VERSION : 1.8
// Fehlerliste:
// Nr.(HEX)     Bedeutung:          
// -------------------------------------------------------------------------------
//  00          Kein Fehler
//  01          Lesen/ Schreiben nicht möglich, kein Codeträger im Bereich des 
//              Schreib-/ Lesekopfes
//  02          Fehler beim Lesen
//  03          Codeträger wurde während des Lesens aus dem Bereich des Schreib-/
//              Lesekopfes entfernt
//  04          Fehler beim Schreiben
//  05          Codeträger wurde während des Schreibens aus dem Bereich des
//              Schreib-/ Lesekopfes entfernt
//  06          Zugriffsfehler auf den Speicher
//  07          AV-Bit gesetzt, aber Befehlskennung fehlt oder ist ungültig.
//              oder: Anzahl Byte ist 00
//  09          Kabelbruch Schreib-/ Lesekopf oder Kopf nicht angeschlossen
//  0F          Inhalt der 1. und 2. Bitleiste sind ungleich
//  10          Startadresse + Anzahl byte > Speicherbereich in Initialisierung
//              angegeben
//  11          Ungültige max. Anzahl Schreibzyklen in Initialisierung angegeben
//  12          Ungültige Speichergröße in Initialisierung angegeben
//  13          Ungültige Größe des Speicherbereichs in Initialisierung angegeben
//  14          Ungültige max. Anzahl Schreibzyklen
//  15          Falscher Codeträger-Typ in Initialisierung angegeben
//  16          Max. Anzahl von 2 kByte überschritten
//  17          Codeträger falsch initialisiert (Vergleich mit Vorgabedaten über
//              Befehlskennung 09 Hex bringt keine Übereinstimmung
//  18          Codeträger noch nicht initialisiert. Alle Byte sind noch 00 Hex
//  30          Überwachungszeit abgelaufen
//  31          ungültiger Auftrag
//  32          Initialisierungsdaten im Instanz-DB für Speicheroptimierung
//              (DBB 178 - DBB 182) nicht korrekt.
   VAR_INPUT
      Init : Bool;   // Neuanlauf der SPS
      Start : Bool;   // Funktion starten
      Reset : Bool;   // FB und Auswerteeinheit BIS-C602-... rücksetzen
      CTTP : Bool;   // Codeträgertyp (0=32Byte;1=64Byte)
      Dynamik : Bool;   // Dynamikbetrieb
      EA_Anfang : Int;   // Anfangsadresse des E/A-Bereiches
      EA_Laenge : Int;   // Länge des E/A-Bereiches
      Auftrag : Int;   // 1=Lesen;2=Schreiben
      DB_Send : Int;   // Datenbaustein für Sendedaten
      Adr_Send : Int;   // Anfangsadresse für Sendedaten
      DB_Empf : Int;   // Datenbaustein für Empfangsdaten
      Adr_Empf : Int;   // Anfangsadresse für Empfangsdaten
      Adr_Traeger : Int;   // Anfangsadresse im Codeträger
      Laenge_Traeger : Int;   // Datenlaenge im Codeträger
      Ueberwzeit : S5Time;   // Überwachungszeit für Senden und Empfangen
      UWZ_Timer : Timer;   // Timer für Überwachungszeit
   END_VAR
   VAR_OUTPUT
      Fertig : Bool;   // Fertig-Bit, Auftrag beendet
      Fehler : Bool;   // Auftrag mit Fehler beendet
      FehlerNr : Int;   // Fehlernummer
      Dig_In : Bool;   // Status des Digitaleingangs an der Auswerteeinheit
      CT_Vorhanden : Bool;   // Codetag vorhanden und Daten im Eingangspuffer gültig
   END_VAR
   VAR
      ZeigerByte : Int;   // Aktuelle Lese-/ Schreibadresse
      LaengeByte : Int;   // Anzahl Byte für Lese-/ Schreibzyklus
      ByteProSeite : Int;   // Anzahl maximaler Nutzbyte pro Seite
      Gesamtbyte : Int;   // Gesamtbyte die gelesen bzw. geschrieben werden
      LesenAktiv : Bool;   // Funktion Lesen ist aktiv
      SchreibenAktiv : Bool;   // Funktion Schreiben ist aktiv
      ResetAktiv : Bool;   // Funktion rücksetzen ist aktiv
      Toggle : Bool;   // Letzer Zustand des Toggle-Bit
      ErsterZyklus : Bool;   // Erster Schreib-/ Lesezyklus
      FP_Start : Bool;   // Flankenmerker Start
      IMP_Start : Bool;   // Impulsmerker Start
      FP_Reset : Bool;   // Flankenmerker Reset
      IMP_Reset : Bool;   // Impulsmerker Reset
      FP_CTPR : Bool;   // Flankenmerker Codetag-Present
      IMP_CTPR : Bool;   // Impulsmerker Codetag-Present
      InitSpOpAktiv : Bool;   // Funktion Init Speicheroptimierung
      stat8 : Int;
      SeiteEingang : Array[0..127] of Byte;
      SeiteAusgang : Array[0..6] of Byte;
      Nr_1_Speicherbereich : Byte;   // Nummer des 1. Speicherbereichs
      CT_Speichergroesse : Byte;   // Speichergröße des Codeträger
      Anz_Schreibzyklen : Byte;   // zulässige Anzahl Schreibzyklen
      Anz_byte_high : Byte;   // Max. Anzahl Byte je Zyklus High-byte
      Anz_byte_low : Byte;   // Max. Anzahl Byte je Zyklus Low-Byte
      Init_Fe : Bool;   // Initialisierung Speicheroptimierung
      Offset : DInt;   // Instanz-DB Offset
      OffsetEin : DInt;   // Offset Eingangsarray
      OffsetAus : DInt;   // Offset Ausgangsarray
   END_VAR
   VAR_TEMP
      InstanzDB : Int;   // Instanz-DB Nummer
      LOG_1 : Bool;   // Logisch 1
      Sp_start : Bool;   // Bei Fehler wird hier der Flankenmerker Start zwischengespeichert
      temp : Byte;   // Temporäre Variable
      schleife : Int;   // Schleifenzähler
      DB_Empf1 : Int;
      DB_Send1 : Int;
      DB_Init1 : Int;
   END_VAR
BEGIN

REGION Network 1: SPS Anlauf
   // Initialisierung Instanz-Bereich
         AN    #LOG_1;
         S     #LOG_1;

         TAR2;  // Bit-Offset des Instanz-DB
         SLD   8;
         SRD   8;
         L     8;
         /D;  // Offset Instanz-DB
         T     #Offset;
         L     42;
         +I;
         T     #OffsetEin;  // Offset des Eingangsarray
         L     #Offset;
         L     170;
         +I;
         T     #OffsetAus;  // Offset des Ausgangsarray
         L     #Offset;
         SLD   3;
         LAR1;

         AN    #Init;
         JC    M002;
         L     0;
         T     DID[AR1, P#30.0];  //DID30
         T     DID[AR1, P#34.0];  //DID34
         T     DID[AR1, P#38.0];  //DID38
         T     #FehlerNr;
         S     #Fertig;
         R     #Fehler;
         R     #Init_Fe;
         R     #UWZ_Timer;
         BEU;
END_REGION

REGION Network 2: Eingangsdaten einlesen in Empfangs-DB
   // Bitleiste 1 einlesen in Instanz-DB
   M002: L     #EA_Anfang;
         SLD   3;
         LAR1;  // Adresse Bitleiste 1 Pointerformat
         L     PIB[AR1, P#0.0];  // Bitleiste 1 einlesen
         T     #temp;
         L     #OffsetEin;  // Anfangsadresse 1. Bitleiste im Instanz-DB
         SLD   3;
         LAR1;
         L     #temp;
         T     DIB[AR1, P#0.0];  // Bitleiste 1 in Instanz-DB schreiben
   // Bitleiste 2 einlesen in Instanz-DB
         L     #EA_Anfang;
         L     #EA_Laenge;
         +I;
         L     1;
         -I;
         SLD   3;
         LAR1;  // Adresse Bitleiste 2 Pointerformat
         L     PIB[AR1, P#0.0];  // Bitleiste 2 einlesen
         T     #temp;
         L     #OffsetEin;
         L     1;
         -I;
         L     #EA_Laenge;  // Anfangsadresse 2. Bitleiste im Instanz-DB
         +I;
         SLD   3;
         LAR1;
         L     #temp;
         T     DIB[AR1, P#0.0];  // Bitleiste 2 in Instanz-DB schreiben
         L     #OffsetEin;
         SLD   3;
         LAR1;
         L     DIB[AR1, P#0.0];  //DIB42 Bitleiste 1
         L     #temp;
         <>I;
         BEC;  // Bitleisten unterschiedlich -> BEB
   // Fehlermeldungen abfragen
         AN    DIX[AR1, P#0.3];  //DIX42.3 Fehler vorhanden ?
         O     #Reset;  // oder Reset
         JC    wt1;
         L     #EA_Anfang;
         L     1;
         +I;
         SLD   3;
         LAR1;
         L     PIB[AR1, P#0.0];  // Fehlernummer laden
         T     #FehlerNr;
         A     #LOG_1;
         JU    Fehe;
   //
   wt1:  L     #OffsetEin;
         SLD   3;
         LAR1;
         A     DIX[AR1, P#0.4];  //DIX42.4
         =     #Dig_In;
   // Eingangsdaten direkt in Instanz-DB einlesen
         A     DIX[AR1, P#0.0];  //DIX42.0 Codetag present
         FP    #FP_CTPR;
         =     #IMP_CTPR;
         AN    #IMP_CTPR;  // Wenn keine pos. Flanke CT_Present, dann Sprung
         JC    wt2;
         L     1;
         T     #schleife;  // Schleifenzähler vorbelegen
   lp1:  L     #schleife;
         L     #EA_Anfang;
         +I;
         SLD   3;
         LAR1;  // aktuelle einzulesende E-Adresse im Pointerformat
         L     PIB[AR1, P#0.0];  // Eingangsbyte indirekt einlesen
         T     #temp;
         L     #OffsetEin;
         L     #schleife;
         +I;
         SLD   3;
         LAR1;  // aktuelle Schreibadresse im Instanz-DB
         L     #temp;
         T     DIB[AR1, P#0.0];  // akt. Eingangsbyte schreiben in Instanz-DB
         L     #schleife;
         L     1;
         +I;
         T     #schleife;  // Schleifenzähler um 1 erhöhen
         L     #EA_Laenge;
         L     2;
         -I;
         L     #schleife;
         >=I;
         JC    lp1;
         A     #LOG_1;
         =     #CT_Vorhanden;
         JU    wt3;
   wt2:  L     #OffsetEin;
         SLD   3;
         LAR1;
         AN    DIX[AR1, P#0.0];  //DIX42.0 Wenn Kein CT_Present vom BIS
         R     #CT_Vorhanden;
   wt3:  NOP   0;
END_REGION

REGION Network 3: Auswerteeinheit rücksetzten
         O     #Reset;  // FB-Eingang Reset
         FP    #FP_Reset;  // Hilfsmerker positive Flanke
         =     #IMP_Reset;  // Impulsmerker, ist einen Zyklus "1"
         A     #IMP_Reset;
         S     #ResetAktiv;
         AN    #ResetAktiv;
         JC    M014;
         R     #LesenAktiv;
         R     #SchreibenAktiv;
         R     #InitSpOpAktiv;
         R     #Toggle;
         R     #Fehler;
         R     #Init_Fe;
         L     0;
         T     #ZeigerByte;
         T     #Gesamtbyte;
         T     #FehlerNr;
         L     #OffsetEin;
         SLD   3;
         LAR1;
         AN    DIX[AR1, P#0.7];  //DIX42.7 Betriebsbereit BIS
         JC    M013;
         L     #OffsetAus;  // Offset Ausgangsarrey
         SLD   3;
         LAR1;
         L     0;
         T     DIB[AR1, P#0.0];  //DIB170 Bitleiste rücksetzen
         S     DIX[AR1, P#0.2];  //DIX170.2 Resetbit setzen
         JU    M012;
   M013: L     #OffsetAus;
         SLD   3;
         LAR1;
         L     0;
         T     DIB[AR1, P#0.0];  //DIB170 Bitleiste rücksetzen
         R     #ResetAktiv;  // Rücksetzen beendet
   M012: L     DIB[AR1, P#0.0];  //DIB170
         T     #temp;
         L     #EA_Anfang;  //1. Bitleiste an Ausgangsbyte übergeben
         SLD   3;
         LAR1;
         L     #temp;
         T     PQB[AR1, P#0.0];
         L     #EA_Anfang;  // Adresse 2. Bitleiste
         L     #EA_Laenge;
         +I;
         L     1;
         -I;
         SLD   3;
         LAR1;
         L     #temp;
         T     PQB[AR1, P#0.0];
   M014: NOP   0;
END_REGION

REGION Network 4: Startauslösung?
         L     #OffsetEin;
         SLD   3;
         LAR1;
         AN    DIX[AR1, P#0.6];  //DIX42.6 Head Fehler
         JC    star;
         O     #ResetAktiv;
         O     #Reset;
         JC    M020;
         L     #stat8;  // Zähler um Kabelbruch nicht sofort
         +     1;  // wirksam werden zu lassen.
         T     #stat8;
         L     30;
         <>I;
         JC    M020;
         L     #stat8;  // Zähler um Kabelbruch nicht sofort
         +     -1;  // wirksam werden zu lassen.
         T     #stat8;
         L     9;
         JU    Fehl;
   star: L     0;
         T     #stat8;
         AN    #SchreibenAktiv;
         AN    #LesenAktiv;
         AN    #InitSpOpAktiv;
         AN    #ResetAktiv;
         AN    DIX[AR1, P#0.1];  //DIX42.1 Auftrag erkannt und begonnen
         AN    DIX[AR1, P#0.3];  //DIX42.3 Auftrag fehlerhaft/ abgebrochen
         A     DIX[AR1, P#0.7];  //DIX42.7 BIS betriebsbereit
         =     #Fertig;
         A     #Start;  // FB-Eingang Start
         FP    #FP_Start;  // Hilfsmerker positive Flanke
         =     #IMP_Start;  // Impulsmerker, ist einen Zyklus "1"

         A(;
         O     #IMP_Start;  // Überwachungszeit starten
         O     DIX[AR1, P#0.1];  //DIX42.1 Auftrag angenommen
         );
         AN    DIX[AR1, P#0.3];  //DIX42.3
         AN    #Dynamik;
         AN    #Init_Fe;
         L     #Ueberwzeit;
         SD    #UWZ_Timer;
         AN    #UWZ_Timer;
         JC    M020;
         L     48;  // Überwachungszeit abgelaufen
         JU    Fehl;
   M020: AN    #LesenAktiv;
         AN    #SchreibenAktiv;
         AN    #InitSpOpAktiv;
         A(;
         AN    #IMP_Start;
         ON    #Fertig;
         O     DIX[AR1, P#0.1];  //DIX42.1
         );
         BEC;
END_REGION

REGION Network 5: Initialisieren
         O     #LesenAktiv;
         JC    Lese;
         O     #SchreibenAktiv;
         JC    Schr;
         O     #InitSpOpAktiv;  //Speicheroptimierung initialisieren
         JC    Init;
         R     #Fehler;
         R     #Init_Fe;
         L     #OffsetAus;
         SLD   3;
         LAR1;
         L     0;
         T     #FehlerNr;
         T     DIB[AR1, P#0.0];  //DIB170 1. Bitleiste rücksetzen
         A     #CTTP;
         =     DIX[AR1, P#0.7];  //DIX170.7 Codeträgertyp parametrieren
         A     #LOG_1;
         S     DIX[AR1, P#0.0];  //DIX170.0 Auftrag vorhanden setzten
   // Leseauftrag?
         L     #Auftrag;  // Auftragsnummer laden
         L     1;
         <>I;
         JC    M025;
         S     #LesenAktiv;  // gleich "1" -> Leseauftrag
         L     1;
         T     DIB[AR1, P#1.0];  //DIB171
         L     #Adr_Empf;
         T     #ZeigerByte;
         JU    M035;
   // Schreibauftrag?
   M025: L     #Auftrag;  // Auftragsnummer laden
         L     2;
         <>I;
         JC    M026;
         S     #SchreibenAktiv;  // gleich "2" -> Schreibauftrag
         L     2;
         T     DIB[AR1, P#1.0];  //DIB171
         L     #Adr_Send;
         T     #ZeigerByte;
         JU    M035;
   //CT Initialisieren, Speicheroptimiert?
   // CT initialisieren
   M026: L     #Auftrag;
         L     8;
         <>I;
         JC    M027;
         L     8;
         T     DIB[AR1, P#1.0];  //DIB171
         L     178;
         L     #Offset;
         +I;
         T     #ZeigerByte;
         L     0;
         T     DIB[AR1, P#8.0];  //DIB178 Datum Nummer 1. Speicherbereich
         L     5;  // 5 Byte Initdaten
         T     #LaengeByte;
         JU    M028;
   // Flash initialisieren, Init-Überwachung
   M027: L     #Auftrag;
         L     9;
         <>I;
         JC    M030;
         L     9;
         T     DIB[AR1, P#1.0];  //DIB171
         L     179;
         L     #Offset;
         +I;
         T     #ZeigerByte;
         L     0;  // keine weiteren Daten mehr
         T     #LaengeByte;
   M028: S     #InitSpOpAktiv;
         JU    Go;
   M030: L     49;  // ungültiger Auftrag
         JU    Fehl;
   // Initialisierungswerte überprüfen
   Go:   L     1;  // Wert 01 Hex
         L     DIB[AR1, P#9.0];  //DIB179 Datum CT-Größe
         >I;
         JC    InFe;
         L     13;  // Wert 0D Hex
         >I;
         JC    InFe;
         L     1;  // Wert 01 Hex
         L     DIB[AR1, P#10.0];  //DIB180 Datum Anzahl Schreibzyklen
         >I;
         JC    InFe;
         L     10;  // Wert 0A Hex
         ==I;
         JC    In2;
         TAK;
         L     5;  //Wert 05 Hex
         >I;
         JC    InFe;
   In2:  L     DIW[AR1, P#11.0];  //DIW181 max. Anzahl Byte Schreib-/Lesezyklen
         L     4096;  // Wert 1000 Hex
         <=D;
         JC    M035;
   InFe: A     #LOG_1;
         S     #Init_Fe;
         L     50;  // Falsche Init-Daten
         JU    Fehl;
   // Erster Zyklus
   M035: AN    #ErsterZyklus;
         S     #ErsterZyklus;
         R     #Fertig;
   // Berechnungen
         L     #EA_Laenge;
         L     2;  // 2 Bitleisten
         -I;
         T     #ByteProSeite;  // Nutzdaten pro Seite

         L     #Laenge_Traeger;
         T     #Gesamtbyte;
END_REGION

REGION Network 6: Auftrag senden
   // Die erste Bitleiste wird gespiegelt. Auftrag (Lesen, Schreiben) wird 
   // gesendet.
   // Befehlsanhang generieren
         L     #Adr_Traeger;  // Anfang des Datenträgers laden
         CAW;  // Low- und Highbyte tauschen
         AN    #InitSpOpAktiv;  // Initialisieren nicht anktiv
         JC    BHG1;
         L     DIW[AR1, P#9.0];  //DIW179 2. und 3. Initbyte
   BHG1: T     DIW[AR1, P#2.0];  //DIW172 ins 2. und 3. Byte des Ausgangspuffers schreiben
         L     #Laenge_Traeger;  // Laenge des Datenträgers laden
         CAW;  // Low- und Highbyte tauschen
         AN    #InitSpOpAktiv;  // Initialisieren nicht anktiv
         JC    BHG2;
         L     DIW[AR1, P#11.0];  //DIW181 4. und 5. Initbyte
   BHG2: T     DIW[AR1, P#4.0];  //DIW174 ins 4. und 5. Byte des Ausgangspuffers schreiben

   // Erste Bitleiste spiegeln auf letztes Byte
         L     #OffsetAus;
         SLD   3;
         LAR1;
         L     DIB[AR1, P#0.0];  // Bitleiste 1
         T     #temp;
         L     #Offset;
         L     176;  // Adresse 2. Bitleiste
         +I;
         SLD   3;
         LAR1;
         L     #temp;  // 1.Bitleiste kopieren auf 2. Bitleiste
         T     DIB[AR1, P#0.0];
   //    Auftrag schreiben
         L     0;
         T     #schleife;  // Schleifenzähler rücksetzen
   lp2:  L     #OffsetAus;
         L     #schleife;
         +I;
         SLD   3;
         LAR1;  // aktuelle Quelladresse
         L     DIB[AR1, P#0.0];
         T     #temp;
         L     #EA_Anfang;
         L     #schleife;
         +I;
         SLD   3;
         LAR1;  // aktuelle Zieladresse
         L     #temp;
         T     PQB[AR1, P#0.0];
         L     #schleife;
         L     1;
         +I;
         T     #schleife;
         L     6;
         <I;
         JC    lp2;  // 1. Bitleiste + Auftrag senden
         L     #OffsetAus;
         SLD   3;
         LAR1;
         L     DIB[AR1, P#0.0];  //DIB 170
         T     #temp;
         L     #EA_Anfang;
         L     #EA_Laenge;
         +I;
         L     1;
         -I;
         SLD   3;
         LAR1;  // Adresse 2. Bitleiste im Pointerformat
         L     #temp;
         T     PQB[AR1, P#0.0];  // 2. Bitleiste senden
         BEU;
END_REGION

REGION Network 7: Lesen
   Lese: L     #OffsetEin;
         SLD   3;
         LAR1;
         ON    DIX[AR1, P#0.2];  //DIX42.2 Auftrag beendet
         O     DIX[AR1, P#0.3];  //DIX42.3
         BEC;
         AN    #ErsterZyklus;
         A(;
         A     #Toggle;  // Toggle-Zustand letzter Zyklus
         A     DIX[AR1, P#0.5];  //DIX42.5 Aktuelles Toggle-Bit
         O;
         AN    #Toggle;  // Toggle-Zustand letzter Zyklus
         AN    DIX[AR1, P#0.5];  //DIX42.5 Aktuelles Toggle-Bit
         );
         BEC;

         L     #ByteProSeite;
         L     #Gesamtbyte;
         <=I;
         JC    M050;
         T     #LaengeByte;  // Nutzdaten kleiner Nutzdaten pro Seite
         JU    M055;
   M050: L     #ByteProSeite;
         T     #LaengeByte;  // Nutzdaten größer gleich Nutzdaten pro Seite
   M055: L     #DB_Empf;
         T     #DB_Empf1;
         OPN   DB[ #DB_Empf1];
         L     0;
         T     #schleife;  // Schleifenzähler rücksetzen
   lp3:  L     #schleife;
         L     #EA_Anfang;
         +I;
         L     1;
         +I;
         SLD   3;
         LAR1;  // Leseadresse Eingang im Pointerformat
         L     PIB[AR1, P#0.0];
         T     #temp;
         L     #ZeigerByte;
         L     #schleife;
         +I;
         SLD   3;
         LAR1;  // Zieladresse Empfangs-DB im Pointerformat
         L     #temp;
         T     DBB[AR1, P#0.0];
         L     #schleife;
         L     1;
         +I;
         T     #schleife;
         L     #LaengeByte;
         <I;
         JC    lp3;
         JU    M070;
END_REGION

REGION Network 8: Schreiben
   Schr: A     DIX[AR1, P#0.2];  //DIX42.2 Auftrag beendet
         JC    M080;
         ON    DIX[AR1, P#0.1];  //DIX42.1 Auftrag begonnen
         O     DIX[AR1, P#0.3];  //DIX42.3 Auftrag Fehler
         BEC;
         A(;
         A     #Toggle;  // Toggle-Zustand letzter Zyklus
         A     DIX[AR1, P#0.5];  //DIX42.5 Aktuelles Toggle-Bit
         O;
         AN    #Toggle;  // Toggle-Zustand letzter Zyklus
         AN    DIX[AR1, P#0.5];  //DIX42.5 Aktuelles Toggle-Bit
         );
         BEC;

         L     #ByteProSeite;
         L     #Gesamtbyte;
         <=I;
         JC    M150;
         T     #LaengeByte;  // Nutzdaten kleiner Nutzdaten pro Seite
         JU    M155;
   M150: L     #ByteProSeite;
         T     #LaengeByte;  // Nutzdaten größer gleich Nutzdaten pro Seite
   //Nutzdaten in Ziel-DB uebertragen
   M155: L     #DB_Send;
         T     #DB_Send1;
         OPN   DB[ #DB_Send1];
         L     0;
         T     #schleife;
   lp5:  L     #ZeigerByte;
         L     #schleife;
         +I;
         SLD   3;
         LAR1;
         L     DBB[AR1, P#0.0];
         T     #temp;
         L     #EA_Anfang;
         L     1;
         +I;
         L     #schleife;
         +I;
         SLD   3;
         LAR1;
         L     #temp;
         T     PQB[AR1, P#0.0];
         L     #schleife;
         L     1;
         +I;
         T     #schleife;
         L     #LaengeByte;
         <I;
         JC    lp5;
         JU    M070;
END_REGION

REGION Network 9: CT Initialisieren, Speicheroptimiert
   Init: L     #OffsetEin;
         SLD   3;
         LAR1;
         A     DIX[AR1, P#0.2];  //DIX42.2 Auftrag beendet
         JC    M080;
         ON    DIX[AR1, P#0.1];  //DIX42.1 Auftrag begonnen
         O     DIX[AR1, P#0.3];  //DIX42.3 Auftrag Fehler
         BEC;
         A(;
         A     #Toggle;  // Toggle-Zustand letzter Zyklus
         A     DIX[AR1, P#0.5];  //DIX42.5 Aktuelles Toggle-Bit
         O;
         AN    #Toggle;  // Toggle-Zustand letzter Zyklus
         AN    DIX[AR1, P#0.5];  //DIX42.5 Aktuelles Toggle-Bit
         );
         BEC;

         L     0;
         T     #schleife;
   lp7:  L     #ZeigerByte;
         L     #schleife;
         +I;
         SLD   3;
         LAR1;
         L     DIB[AR1, P#0.0];
         T     #temp;
         L     #EA_Anfang;
         L     1;
         +I;
         L     #schleife;
         +I;
         SLD   3;
         LAR1;
         L     #temp;
         T     PQB[AR1, P#0.0];
         L     #schleife;
         L     1;
         +I;
         T     #schleife;
         L     #LaengeByte;
         <I;
         JC    lp7;
END_REGION

REGION Network 10: schreiben/ lesen
   M070: L     #OffsetEin;
         SLD   3;
         LAR1;
         L     #Gesamtbyte;  //Bytes die noch uebertragen werden müssen
         L     #LaengeByte;  //Bytes die in diesem Zyklus uebertragen wurden
         -I;  //Bytes hinzuaddieren
         T     #Gesamtbyte;

         L     #ZeigerByte;  // Zielbyte erhöhen um Nutzdatenlaenge des E/A-Bereichs
         L     #LaengeByte;
         +I;
         T     #ZeigerByte;


         A     DIX[AR1, P#0.5];  //DIX42.5
         =     #Toggle;  // Toggle-Zustand speichern
         L     #OffsetAus;
         SLD   3;
         LAR1;
         AN    DIX[AR1, P#0.6];
         =     DIX[AR1, P#0.6];  // Toggle-Bit invertieren im Instanz-DB 1. Bitleiste
         L     DIB[AR1, P#0.0];  //DIB170
         T     DIB[AR1, P#6.0];  //DIB176 Bitleiste 1 kopieren in Bitleiste 2
         T     #temp;

         L     #EA_Anfang;
         SLD   3;
         LAR1;
         L     #temp;
         T     PQB[AR1, P#0.0];  //  1. Bitleiste aus Instanz-DB übertragen auf Ausgang

         L     #EA_Anfang;
         L     #EA_Laenge;
         +I;
         L     1;
         -I;
         SLD   3;
         LAR1;
         L     #temp;
         T     PQB[AR1, P#0.0];  //  2. Bitleiste aus Instanz-DB übertragen auf Ausgang

         A     #ErsterZyklus;
         R     #ErsterZyklus;

         L     #Gesamtbyte;
         L     0;
         >D;
         BEC;  // Übertragung noch nicht beendet
   M080: L     #OffsetEin;
         SLD   3;
         LAR1;
         AN    DIX[AR1, P#0.2];  //DIX42.2
         BEC;
   m090: L     #OffsetAus;
         SLD   3;
         LAR1;
         A     #LOG_1;
         R     #LesenAktiv;
         R     #SchreibenAktiv;
         R     #InitSpOpAktiv;
         R     #Toggle;
         R     DIX[AR1, P#0.0];  //DIX170.0 Auftrag vorhanden rücksetzten

         L     #EA_Anfang;  // Auftrag vorhanden rücksetzen 1. Bitleiste
         SLD   3;
         LAR1;
         L     0;
         T     PQB[AR1, P#0.0];

         L     #EA_Anfang;  // Auftrag vorhanden rücksetzen 2. Bitleiste
         L     #EA_Laenge;
         +I;
         L     1;
         -I;
         SLD   3;
         LAR1;
         L     0;
         T     PQB[AR1, P#0.0];
         BEU;
END_REGION

REGION Network 11: Fehler eintragen
   Fehl: T     #FehlerNr;
   Fehe: L     #Offset;
         SLD   3;
         LAR1;
         S     #Fehler;
         R     #Fertig;
         A     #FP_Start;
         =     #Sp_start;
         L     0;
         T     DID[AR1, P#30.0];  //DID30
         T     DID[AR1, P#34.0];  //DIB34
         T     DID[AR1, P#38.0];  //DIB38
         A     #Sp_start;
         =     #FP_Start;
         JU    m090;
END_REGION
END_FUNCTION_BLOCK

FUNCTION_BLOCK "FB100_Common_Aggregates_General"   // FB100, STL
{ S7_Optimized_Access := 'FALSE' }
VERSION : 0.1
BEGIN

REGION Network 1: These tank is exist
         L     "DB790_PlantParameter".AmountTank;
         JL    nTank;
         JU    Tank00;  // case 0     0 Daytanks selected
         JU    Tank01;  // case 1     1 Daytank selected
         JU    Tank02;  // case 2     2 Daytanks selected
         JU    Tank03;  // case 3     3 Daytanks selected
         JU    Tank04;  // case 4     4 Daytanks selected
         JU    Tank05;  // case 5     5 Daytanks selected
         JU    Tank06;  // case 6     6 Daytanks selected
         JU    Tank07;  // case 7     7 Daytanks selected
         JU    Tank08;  // case 8     8 Daytanks selected
         JU    Tank09;  // case 9     9 Daytanks selected
         JU    Tank10;  // case 10    10 Daytanks selected
         JU    Tank11;  // case 11    11 Daytanks selected
         JU    Tank12;  // case 12    12 Daytanks selected
   //-----
   nTank:NOP   0;
         JU    End;
   //-----
   Tank00:NOP   0;
         SET;
         R     "DB702_Tank_Value".Tank[1].Existing;
         R     "DB702_Tank_Value".Tank[2].Existing;
         R     "DB702_Tank_Value".Tank[3].Existing;
         R     "DB702_Tank_Value".Tank[4].Existing;
         R     "DB702_Tank_Value".Tank[5].Existing;
         R     "DB702_Tank_Value".Tank[6].Existing;
         R     "DB702_Tank_Value".Tank[7].Existing;
         R     "DB702_Tank_Value".Tank[8].Existing;
         R     "DB702_Tank_Value".Tank[9].Existing;
         R     "DB702_Tank_Value".Tank[10].Existing;
         R     "DB702_Tank_Value".Tank[11].Existing;
         R     "DB702_Tank_Value".Tank[12].Existing;
         JU    End;
   //-----
   Tank01:NOP   0;
         SET;
         R     "DB702_Tank_Value".Tank[2].Existing;
         R     "DB702_Tank_Value".Tank[3].Existing;
         R     "DB702_Tank_Value".Tank[4].Existing;
         R     "DB702_Tank_Value".Tank[5].Existing;
         R     "DB702_Tank_Value".Tank[6].Existing;
         R     "DB702_Tank_Value".Tank[7].Existing;
         R     "DB702_Tank_Value".Tank[8].Existing;
         R     "DB702_Tank_Value".Tank[9].Existing;
         R     "DB702_Tank_Value".Tank[10].Existing;
         R     "DB702_Tank_Value".Tank[11].Existing;
         R     "DB702_Tank_Value".Tank[12].Existing;
         JU    End;
   //-----
   Tank02:NOP   0;
         SET;
         R     "DB702_Tank_Value".Tank[3].Existing;
         R     "DB702_Tank_Value".Tank[4].Existing;
         R     "DB702_Tank_Value".Tank[5].Existing;
         R     "DB702_Tank_Value".Tank[6].Existing;
         R     "DB702_Tank_Value".Tank[7].Existing;
         R     "DB702_Tank_Value".Tank[8].Existing;
         R     "DB702_Tank_Value".Tank[9].Existing;
         R     "DB702_Tank_Value".Tank[10].Existing;
         R     "DB702_Tank_Value".Tank[11].Existing;
         R     "DB702_Tank_Value".Tank[12].Existing;
         JU    End;
   //-----
   Tank03:NOP   0;
         SET;
         R     "DB702_Tank_Value".Tank[4].Existing;
         R     "DB702_Tank_Value".Tank[5].Existing;
         R     "DB702_Tank_Value".Tank[6].Existing;
         R     "DB702_Tank_Value".Tank[7].Existing;
         R     "DB702_Tank_Value".Tank[8].Existing;
         R     "DB702_Tank_Value".Tank[9].Existing;
         R     "DB702_Tank_Value".Tank[10].Existing;
         R     "DB702_Tank_Value".Tank[11].Existing;
         R     "DB702_Tank_Value".Tank[12].Existing;
         JU    End;
   //-----
   Tank04:NOP   0;
         SET;
         R     "DB702_Tank_Value".Tank[5].Existing;
         R     "DB702_Tank_Value".Tank[6].Existing;
         R     "DB702_Tank_Value".Tank[7].Existing;
         R     "DB702_Tank_Value".Tank[8].Existing;
         R     "DB702_Tank_Value".Tank[9].Existing;
         R     "DB702_Tank_Value".Tank[10].Existing;
         R     "DB702_Tank_Value".Tank[11].Existing;
         R     "DB702_Tank_Value".Tank[12].Existing;
         JU    End;
   //-----
   Tank05:NOP   0;
         SET;
         R     "DB702_Tank_Value".Tank[6].Existing;
         R     "DB702_Tank_Value".Tank[7].Existing;
         R     "DB702_Tank_Value".Tank[8].Existing;
         R     "DB702_Tank_Value".Tank[9].Existing;
         R     "DB702_Tank_Value".Tank[10].Existing;
         R     "DB702_Tank_Value".Tank[11].Existing;
         R     "DB702_Tank_Value".Tank[12].Existing;
         JU    End;
   //-----
   Tank06:NOP   0;
         SET;
         R     "DB702_Tank_Value".Tank[7].Existing;
         R     "DB702_Tank_Value".Tank[8].Existing;
         R     "DB702_Tank_Value".Tank[9].Existing;
         R     "DB702_Tank_Value".Tank[10].Existing;
         R     "DB702_Tank_Value".Tank[11].Existing;
         R     "DB702_Tank_Value".Tank[12].Existing;
         JU    End;
   //-----
   Tank07:NOP   0;
         SET;
         R     "DB702_Tank_Value".Tank[8].Existing;
         R     "DB702_Tank_Value".Tank[9].Existing;
         R     "DB702_Tank_Value".Tank[10].Existing;
         R     "DB702_Tank_Value".Tank[11].Existing;
         R     "DB702_Tank_Value".Tank[12].Existing;
         JU    End;
   //-----
   Tank08:NOP   0;
         SET;
         R     "DB702_Tank_Value".Tank[9].Existing;
         R     "DB702_Tank_Value".Tank[10].Existing;
         R     "DB702_Tank_Value".Tank[11].Existing;
         R     "DB702_Tank_Value".Tank[12].Existing;
         JU    End;
   //-----
   Tank09:NOP   0;
         SET;
         R     "DB702_Tank_Value".Tank[10].Existing;
         R     "DB702_Tank_Value".Tank[11].Existing;
         R     "DB702_Tank_Value".Tank[12].Existing;
         JU    End;
   //-----
   Tank10:NOP   0;
         SET;
         R     "DB702_Tank_Value".Tank[11].Existing;
         R     "DB702_Tank_Value".Tank[12].Existing;
         JU    End;
   //-----
   Tank11:NOP   0;
         SET;
         R     "DB702_Tank_Value".Tank[12].Existing;
         JU    End;
   //-----
   Tank12:NOP   0;
         JU    End;
   //-----
   End:  NOP   0;
END_REGION
END_FUNCTION_BLOCK

FUNCTION_BLOCK "FB101_Common_Aggregates_C1"   // FB101, STL
TITLE = Agitators,Tanks, Refilling, tempering
{ S7_Optimized_Access := 'FALSE' }
AUTHOR : KT242
VERSION : 0.1
// Common aggregates
   VAR_TEMP
      Real_dummy : Real;
      CompUsedForShot : Array[1..16] of Bool;
      Dummy : Bool;
      MH_open : Bool;
      K_Tanklager : Bool;
      Temp_Vacuum_active : Bool;
      Temp_Cooling : Bool;
      Temp_Pentan_Enabling : Bool;
      Temp_Filling_Enable : Bool;
      Temp_Aggitator_Enable : Bool;
      Temp_BefuellungAngewaehlt : Bool;
      Temp_Filling_Ends : Bool;
      Temp_Filling_Valve : Bool;
      Temp_StartExtern : Bool;
      Temp_WithFillingPump : Bool;
      Temp_FillingPumpActive : Bool;
      Valid_Circulation : Bool;
      temp_V_Barrel_C1 : Bool;
      Temp_FaultGrp3 : Bool;
      Temp_SwitchONTemp : Bool;
      Temp_EnableTempering : Bool;
      Temp_RequestFillAuto : Bool;
      HF_Pulse_alarm : Bool;
      Temp_RetVal_SFC14 : Word;
      Temp_RetVal_SFC15 : Word;
      Temp_SetValue_TG : Int;
      Temp_Refilling_Barrel : Bool;   // Toggle bit, if refilling over barrel station is activated
   END_VAR
BEGIN

REGION Network 1: Toggle bit, if refilling over barrel station is activated
   // Copy Control bits for module to local area
         L;
         LAR1;
         L     "DB619_State_MPart".ShotMa[1].ShotData.Comp_at_Shot;
         L     "DB619_State_MPart".ShotMa[2].ShotData.Comp_at_Shot;
         OD;
         CAW;
         T     LW[AR1, P#0.0];

         A     "DB612_Tank_State".Tank[1].Switch_Refilling_from_Barrel_ON_OFF;
         =     #Temp_Refilling_Barrel;
END_REGION

REGION Network 2: Signal a mixinghead opens
         O     "DB619_State_MPart".Mixinghead[1].Shotcounter."01";
         O     "DB619_State_MPart".Mixinghead[1].Shotcounter."02";
         O     "DB619_State_MPart".Mixinghead[1].Shotcounter."03";
         O     "DB619_State_MPart".Mixinghead[1].Shotcounter."04";
         O     "DB619_State_MPart".Mixinghead[1].Shotcounter."05";
         O     "DB619_State_MPart".Mixinghead[1].Shotcounter."06";
         O     "DB619_State_MPart".Mixinghead[1].Shotcounter."07";
         O     "DB619_State_MPart".Mixinghead[1].Shotcounter."08";
         O     "DB619_State_MPart".Mixinghead[1].Shotcounter."09";
         O     "DB619_State_MPart".Mixinghead[1].Shotcounter."10";
         O     "DB619_State_MPart".Mixinghead[1].Shotcounter."11";
         O     "DB619_State_MPart".Mixinghead[1].Shotcounter."12";
         O     "DB619_State_MPart".Mixinghead[1].Shotcounter."13";
         O     "DB619_State_MPart".Mixinghead[1].Shotcounter."14";
         O     "DB619_State_MPart".Mixinghead[1].Shotcounter."15";
         O     "DB619_State_MPart".Mixinghead[1].Shotcounter."16";
         A     #CompUsedForShot[1];
         =     #MH_open;
END_REGION

REGION Network 3: GBE
         CALL  "FC920_PV_Calc_Act_Value"
         ( IN_Act_Value_read := "DB702_Tank_Value".Tank[1].With_Nucleation,
           IN_Act_Value_ext  := FALSE,
           IN_Ext_Value      := #Real_dummy,
           IN_Read_Double    := FALSE,
           IN_FLT_Needful    := TRUE,
           IN_FLT_Reset      := "DB009_Faults".Faults_Reset_FKT_M1,
           IO_Any_ArrayPV    := "DB602_PV_Tank".Tank[1].Nucleation,
           IO_Fault_Sensor   := "DB822_Error_Tank".Refilling_Tank[1].FLT_NucleationSensor_broken_wire,
           IO_New_Fault      := "DB009_Faults".Faultschanging_M1,
           IO_FLT_Level_3    := "DB009_Faults".Faults_FKT_Grp_3_M1
         );
   //-----
         O     "DB009_Faults".Faults_Reset_FKT_M1;
         ON    "DB702_Tank_Value".Tank[1].With_Nucleation;
         R     "DB822_Error_Tank".Refilling_Tank[1].FLT_supply_nucleation;
         R     "DB822_Error_Tank".Refilling_Tank[1].FLT_nucleation;
   //-
         AN    "F_GBE_C1";
         A     "DB702_Tank_Value".Tank[1].With_Nucleation;
         AN    "DB822_Error_Tank".Refilling_Tank[1].FLT_supply_nucleation;
         S     "DB009_Faults".Faultschanging_M1;
         S     "DB822_Error_Tank".Refilling_Tank[1].FLT_supply_nucleation;
   //-
         A     "F_GBE_Faulty_C1";
         A     "DB702_Tank_Value".Tank[1].With_Nucleation;
         AN    "DB822_Error_Tank".Refilling_Tank[1].FLT_nucleation;
         S     "DB009_Faults".Faultschanging_M1;
         S     "DB822_Error_Tank".Refilling_Tank[1].FLT_nucleation;
   //-
         O     "DB822_Error_Tank".Refilling_Tank[1].FLT_nucleation;
         O     "DB822_Error_Tank".Refilling_Tank[1].FLT_supply_nucleation;
         S     "DB009_Faults".Faults_FKT_Grp_3_M1;
   //-----
END_REGION

REGION Network 4: Filling level
         CALL  "FC920_PV_Calc_Act_Value"
         ( IN_Act_Value_read := "DB702_Tank_Value".Tank[1].With_Level_Probe,
           IN_Act_Value_ext  := FALSE,
           IN_Ext_Value      := #Real_dummy,
           IN_Read_Double    := FALSE,
           IN_FLT_Needful    := TRUE,
           IN_FLT_Reset      := "DB009_Faults".Faults_Reset_FKT_M1,
           IO_Any_ArrayPV    := "DB602_PV_Tank".Tank[1].Level,
           IO_Fault_Sensor   := "DB822_Error_Tank".Refilling_Tank[1].FLT_LevelSensor_broken_wire,
           IO_New_Fault      := "DB009_Faults".Faultschanging_M1,
           IO_FLT_Level_3    := "DB009_Faults".Faults_FKT_Grp_3_M1
         );
   //-----
         AN    "DB702_Tank_Value".Tank[1].DrainTank;
         R     "DB612_Tank_State".Tank[1].Switch_DrainTank_ON_OFF;
   //-----
         CALL  "FC104_FillingSignals"
         ( Tank_exist           := "DB702_Tank_Value".Tank[1].Existing,
           Actual_Level_Value   := "DB602_PV_Tank".Tank[1].Level.PV_ActV.Value,
           IN_With_Level_Probe  := "DB702_Tank_Value".Tank[1].With_Level_Probe,
           IN_With_Triptray     := "DB702_Tank_Value".Tank[1].With_Triptray,
           IN_FLT_Level_Probe   := "DB822_Error_Tank".Refilling_Tank[1].FLT_LevelSensor_broken_wire,
           IN_Max_Level         := "L_DT_max_C1",
           IN_Stop_Fill_Level   := "L_Tank_stop_C1",
           IN_Start_Fill_Level  := "L_Tank_start_C1",
           IN_Min_Level         := "L_Tank_min_C1",
           IN_Triptray          := "L_DripTray_C1",
           IN_DrainTank         := "DB612_Tank_State".Tank[1].Switch_DrainTank_ON_OFF,
           OUT_PreWarnMinLevel  := "DB612_Tank_State".Tank[1].PreWarning_Min_Level,
           OUT_Max_Level        := "DB612_Tank_State".Tank[1].Max_Level,
           OUT_Stop_Fill_Level  := "DB612_Tank_State".Tank[1].Stop_Level_Filling,
           OUT_Start_Fill_Level := "DB612_Tank_State".Tank[1].Start_Level_Filling,
           OUT_Min_Level        := "DB612_Tank_State".Tank[1].Min_Level,
           OUT_Enable_Agitator  := "DB612_Tank_State".Tank[1].Enable_Agitator,
           OUT_Triptray         := "DB612_Tank_State".Tank[1].LevelTriptray,
           IO_TankLevelPar      := "DB702_Tank_Value".Tank[1].TankLevel
         );
   //-----
END_REGION

REGION Network 5: Pentan: Signal machine running to gas warning desk
   //CALL  "FC108_Pentan"
   //         IN_With_Pentan          :="DB702_Tank_Value".Tank[1].With_Filling_Pentane
   //         IN_With_2_Valves        :="DB702_Tank_Value".Tank[1].With_Filling_2Valve
   //         IN_ResetFault           :="DB009_Faults".Faults_Reset_FKT_M1
   //         IN_FirstPLCcycle        :="Flag_Erster_SPS_Zyklus"
   //         IN_OPmode_Valid         :="DB619_State_MPart".Operationmode[1].valid
   //         IN_OPmode_Wekend        :="DB619_State_MPart".Recirculation[1].Weekendswitching
   //         IN_Filling_Selected     :="DB612_Tank_State".Tank[1].Switch_Refilling_ON_OFF
   //         IN_Filling_Start        :="DB612_Tank_State".Tank[1].Filling_Start
   //         IN_Max_Level_Tank       :="DB612_Tank_State".Tank[1].Max_Level
   //         IN_Cycle_runs           :="DB619_State_MPart".Cycle[1].running
   //         IN_Timer_ExhauseSystem  :="TM_ExhauseSystem"
   //         IN_Timer_Overlap_Valves :="TM_Overlap_Valves_Pentan"
   //         IN_Timer_Valve1         :="TM_Valve1_Pentan"
   //         IN_Timer_Valve2         :="TM_Valve2_Pentan"
   //         OUT_EnableComponent     :=#Temp_Pentan_Enabling
   //         OUT_FillingValve1       :="V_ChargingTank_C1"
   //         OUT_FillingValve2       :="V_ChargingTank_C1_2"
   //         IO_Status               :="DB612_Tank_State".Pentan[1]
   //         IO_Fault                :="DB822_Error_Tank".Pentan[1]
   //         IO_NewFault             :="DB009_Faults".Faultschanging_M1
   //         IO_FaultLevel_1         :="DB009_Faults".Faults_FKT_Grp_1_M1
   //         IO_FaultLevel_2         :="DB009_Faults".Faults_FKT_Grp_2_M1
   //         IO_FaultLevel_3         :="DB009_Faults".Faults_FKT_Grp_3_M1
   //-----
   // Signal an GWP, dass die Maschine Kreislauf fahren will
         A     "DB613_Komponent_State".MeteringPump[1].Main_Pumpselection;
         A     "DB619_State_MPart".Recirculation[1].Weekendswitching;
         =     "K_Machine_Running";
   //-----
END_REGION

REGION Network 6: Filling daytank
   //-----
         AN    "DB822_Error_Tank".FeedPump[1].FLT_Dryrunsafety;
         AN    "DB822_Error_Tank".FeedPump[1].FLT_Motorprotection;
         AN    "DB822_Error_Tank".FeedPump[1].FLT_No_Barrel;
         A     "DB619_State_MPart".Operationmode[1].valid;
         A(;
         ON    "DB702_Tank_Value".Tank[1].With_ContainerStation;
         O     "Container_Ready_C1";
         );
         A     #Temp_Pentan_Enabling;
         =     #Temp_Filling_Enable;
   //-----
         A     "Container_Fillpump_run_C1";
         =     #Temp_FillingPumpActive;
   //-----
         A     "DB702_Tank_Value".Tank[1].With_ContainerStation;
         =     #Temp_WithFillingPump;
   //-----
         CALL  "FC102_Refilling"
         ( IN_Selected             := "DB702_Tank_Value".Tank[1].Existing,
           IN_ReleaseRefilling     := "DB619_State_MPart".Operationmode[1].valid,
           IN_FillingPumpActive    := #Temp_FillingPumpActive,
           IN_WithFillingPump      := #Temp_WithFillingPump,
           IN_RecircWeekend        := "DB619_State_MPart".Recirculation[1].Weekendswitching,
           IN_FoamingCycleActive   := "DB619_State_MPart".Cycle[1].running,
           IN_PistonActive         := FALSE,
           IN_MH_is_open           := #MH_open,
           IN_ResetFault           := "DB009_Faults".Faults_Reset_FKT_M1,
           IN_MaxLevelTriptray     := "DB612_Tank_State".Tank[1].LevelTriptray,
           IN_PumpDeselected       := "DB753_MeteringPump".Pump[1].PumpDeselected,
           IN_SetAmountShots       := "DB702_Tank_Value".Tank[1].NoShotFilling,
           IN_PreAgitatingTime     := "DB702_Tank_Value".Tank[1].PreAgitatingTime,
           IN_FillingTimeContr     := "DB702_Tank_Value".Tank[1].FillingTimeControl,
           IN_TimeTillFillingStart := "DB702_Tank_Value".Tank[1].TimeToStartFilling,
           IN_Timer_Refilling      := "TM_Refilling_01",
           OUT_V_Preagitating      := "M_AgitatorBarrel_C1",
           OUT_V_Refilling         := #Temp_Filling_Valve,  // "DB612_Tank_State".Pentan[1].HM_FillingValve // "V_ChargingTank_C1"
           OUT_R_Tankstorage       := #K_Tanklager,
           IO_Status               := "DB612_Tank_State".Tank[1],
           IO_NewFault             := "DB009_Faults".Faultschanging_M1,
           IO_FaultLevel_1         := "DB009_Faults".Faults_FKT_Grp_1_M1,
           IO_FaultLevel_2         := "DB009_Faults".Faults_FKT_Grp_2_M1,
           IO_FaultLevel_3         := "DB009_Faults".Faults_FKT_Grp_3_M1,
           IO_Fault                := "DB822_Error_Tank".Refilling_Tank[1]
         );
   //-----
         A     #Temp_Refilling_Barrel;
         JC    BarrelFill;
         R     "K_Filling_Tank_C1_TL";
         R     "V_ChargingTank_C1_2";

         A     #K_Tanklager;
         A     #Temp_Filling_Valve;
         =     "K_Filling_Tank_C1";
         =     "V_ChargingTank_C1";
         =     "V_Barrel_C1";
         =     "C_Start_Refill_POLY_ON";

         JU    NoBarrelFill;

   BarrelFill:R     "K_Filling_Tank_C1";
         R     "V_ChargingTank_C1";

         A     #K_Tanklager;
         A     #Temp_Filling_Valve;
         =     "K_Filling_Tank_C1_TL";
         =     "V_ChargingTank_C1_2";
         =     "V_Barrel_C1";
         =     "C_Start_Refill_POLY_ON";

   //      U     #Temp_Filling_Enable
   //      U     #Temp_Filling_Valve
   //      =     "DB612_Tank_State".Pentan[1].HM_FillingValve
   //-----
END_REGION

REGION Network 7: Agitator daytank
   //-----
   //-----
   // Das Befüllen soll das Rührwerk nur im Auto ansteuern
   NoBarrelFill:A     "DB612_Tank_State".Tank[1].Fillingtime_runs;
         A     "DB619_State_MPart".Operationmode[1].Auto;
         =     #Temp_RequestFillAuto;

   //      U     #Temp_Pentan_Enabling
   //      U     "DB619_State_MPart".Operationmode[1].valid
   //      UN    "DB823_Error_Metering".MeteringPump[1].FLT_Min_Pressure
   //      UN    "DB822_Error_Tank".Pentan[1].FLT_PreAlam_NitrogenTank
   //      =     #Temp_Aggitator_Enable

   //-----
         CALL  "FC121_Aggitator"
         ( IN_Release               := "DB619_State_MPart".Operationmode[1].valid,  //#Temp_Aggitator_Enable
           IN_ControlVoltage        := "DB619_State_MPart".Operationmode[1].Controllvoltage,
           IN_Reset_fault           := "DB009_Faults".Faults_Reset_FKT_M1,
           IN_Request_Filling       := #Temp_RequestFillAuto,  //"DB612_Tank_State".Tank[1].Fillingtime_runs
           IN_Request_Feed          := 0,
           IN_Request_Cooling       := "DB612_Tank_State".ControllerTankTemp[1].CoolingActive,
           IN_Request_Heating       := "DB612_Tank_State".ControllerTankTemp[1].HeatingActive,
           IN_Fault_Motorprotection := "F_Agitator_C1",
           IN_FaultFreqConverter    := "F_FC_Agitator_C1",
           IN_MaxLevelTray          := "DB612_Tank_State".Tank[1].LevelTriptray,
           IN_EnableLevel           := "DB612_Tank_State".Tank[1].Enable_Agitator,
           IN_TimerDrive            := "TM1_Agitator_01",
           IN_TimerStartUpFConv     := "TM2_Agitator_01",
           IN_Values                := "DB702_Tank_Value".Tank[1].Agitator,
           OUT_MainsContactor       := "M_Agitator_C1",
           OUT_Release_FConverter   := "M_FU_Start_RW_K1",
           IO_Status                := "DB612_Tank_State".Agitator[1],
           IO_NewFault              := "DB009_Faults".Faultschanging_M1,
           IO_FaultLevel_3          := "DB009_Faults".Faults_FKT_Grp_3_M1,
           IO_Faults                := "DB822_Error_Tank".Agitator[1]
         );
END_REGION

REGION Network 8: Tempering Tank Poly
         A     "DB009_Faults".Faults_Reset_FKT_M1;
         R     "DB822_Error_Tank".ControllerTankTemp[1].Fuse_TemperingUnit;
   //-
         AN    "F_Temperiergeraet_C1";
         A     "DB702_Tank_Value".Tank[1].With_Tempering_TempGeraet;
         AN    "DB822_Error_Tank".ControllerTankTemp[1].Fuse_TemperingUnit;
         S     "DB009_Faults".Faultschanging_M1;
         S     "DB822_Error_Tank".ControllerTankTemp[1].Fuse_TemperingUnit;
   //-
         A     "DB822_Error_Tank".ControllerTankTemp[1].Fuse_TemperingUnit;
         S     "DB009_Faults".Faults_FKT_Grp_3_M1;
   //-----
         CALL  "FC920_PV_Calc_Act_Value"
         ( IN_Act_Value_read := TRUE,
           IN_Act_Value_ext  := FALSE,
           IN_Ext_Value      := #Real_dummy,
           IN_Read_Double    := FALSE,
           IN_FLT_Needful    := TRUE,
           IN_FLT_Reset      := "DB009_Faults".Faults_Reset_FKT_M1,
           IO_Any_ArrayPV    := "DB602_PV_Tank".Tank[1].Temp,
           IO_Fault_Sensor   := "DB822_Error_Tank".ControllerTankTemp[1].Sensor_FLT_broken_wire,
           IO_New_Fault      := "DB009_Faults".Faultschanging_M1,
           IO_FLT_Level_3    := "DB009_Faults".Faults_FKT_Grp_3_M1
         );
   //-----
         CALL  "FC916_PV_Limits"
         ( IN_Tolerance_Test     := TRUE,
           IN_Reset_Fault        := "DB009_Faults".Faults_Reset_FKT_M1,
           IO_Any_ArrayPV        := "DB602_PV_Tank".Tank[1].Temp,
           IO_Fault_Warn_upperL  := "DB822_Error_Tank".ControllerTankTemp[1].Warning_limit_plus,
           IO_Fault_Warn_lowerL  := "DB822_Error_Tank".ControllerTankTemp[1].Warning_limit_minus,
           IO_Fault_Alarm_upperL := "DB822_Error_Tank".ControllerTankTemp[1].Alarm_limit_plus,
           IO_Fault_Alarm_lowerL := "DB822_Error_Tank".ControllerTankTemp[1].Alarm_limit_minus,
           IO_New_Fault          := "DB009_Faults".Faultschanging_M1,
           IO_Fault_Level_1      := "DB009_Faults".Faults_FKT_Grp_2_M1,
           IO_Fault_Level_2      := #Dummy,
           IO_Fault_Level_3      := "DB009_Faults".Faults_FKT_Grp_3_M1
         );
   //-----
   //---------------------------------------------
   //  Controller temperature tank poly
   //---------------------------------------------
         O     "DB702_Tank_Value".Tank[1].With_Tempering_VKaltwasser;
         O     "DB702_Tank_Value".Tank[1].With_Tempering_Heizung;
         =     #Temp_EnableTempering;
   //-----
         CALL  "FC105_Tempering"
         ( IN_Exist                := #Temp_EnableTempering,
           IN_Release              := "DB619_State_MPart".Operationmode[1].valid,
           IN_Stop_Tempering       := FALSE,
           IN_F_Fuse               := "F_Heating",
           IN_F_Limit              := FALSE,
           IN_FLT_Ackn             := "DB009_Faults".Faults_Reset_FKT_M1,
           IN_CoolingRequested     := TRUE,
           IN_HeatingRequested     := "DB702_Tank_Value".Tank[1].With_Tempering_Heizung,
           IN_actual_Temp          := "DB602_PV_Tank".Tank[1].Temp.PV_ActV.Value,
           IN_set_Temp             := "DB602_PV_Tank".Tank[1].Temp.PV_SetV.Value,
           Out_act_cooling         := #Temp_Cooling,
           Out_act_request_cooling := #Dummy,
           Out_act_heating         := "K_HeatingTank_C1",
           Out_act_request_heating := #Dummy,
           IO_StateCtrl1           := "DB612_Tank_State".ControllerTankTemp[1],
           IO_ValueCtrl1           := "DB702_Tank_Value".Pt2_Controller[1],
           IO_FaultsCtrl1          := "DB822_Error_Tank".ControllerTankTemp[1],
           IO_NewFault             := "DB009_Faults".Faultschanging_M1,
           IO_FaultLevel_3         := "DB009_Faults".Faults_FKT_Grp_3_M1
         );
   //-----
         A     "DB619_State_MPart".Machine[1].Metering."01";  //Pump running
         A     "DB702_Tank_Value".Tank[1].With_Tempering_WTRL;  // Select from Panel
         A     #Temp_Cooling;
         O(;
         A     "DB613_Komponent_State".HeatexchangerLP[1].CoolingActive;
         A     "DB619_State_MPart".Machine[1].Metering."01";
         A     "DB753_MeteringPump".Pump[1].WithLPHeatExchanger;
         );
         =     "V_Heatexchanger_C1";
   //-----
         ON    "DB619_State_MPart".Machine[1].Metering."01";
         ON    "DB702_Tank_Value".Tank[1].With_Tempering_WTRL;
         A     #Temp_Cooling;
         =     "V_Coolingwater_C1";
   //-----

   // Tempering device gets/sets temperature values with multiplier of 10.
         CALL  CONVERTTO
         ( IN      := "DB602_PV_Tank".Tank[1].Temp.PV_SetV.Value,
           Ret_Val := #Temp_SetValue_TG
         );

         L     #Temp_SetValue_TG;
         L     10;
         *I;
         T     #Temp_SetValue_TG;


         A     "Flag_00_500_Hertz";
         FP    "HF_pulse_alarm_GWK1";
         =     #HF_Pulse_alarm;

   //     CALL  "GWK_PB_TecoCS(CW)e"
   //         IN_With_tempering_unit :="DB702_Tank_Value".Tank[1].With_Tempering_TempGeraet
   //         IN_Flag_alarm          :=#HF_Pulse_alarm
   //         IN_Adr                 :="gwk_temp1~gwk_KRPRO_V6_2_1"
   //         IN_Sl_Akt              :=1
   //         IN_TL_KomF             :=1
   //         IN_On                  :="DB612_Tank_State".ControllerTankTemp[1].Switch_Temp_ON_OFF
   //         IN_Release             :="DB619_State_MPart".Operationmode[1].valid//"DB10_State_MC1".Operating_mode.valid
   //         IN_Weekendmode         :=FALSE
   //         IN_Fault_quit          :="DB009_Faults".Faults_Reset_FKT_M1
   //         IN_Fuse                :="F_Temperiergeraet_C1"
   //         IN_Setvalue            :=#Temp_SetValue_TG
   //         IN_Setvalue_weekend    :=#Temp_SetValue_TG
   //         IN_Actvalue_tool       :="DB602_PV_Tank".Tank[1].Temp.PV_ActV.Value
   //         RetVal_SFC14           :=#Temp_RetVal_SFC14
   //         RetVal_SFC15           :=#Temp_RetVal_SFC15
   //         PBData                 :="DB905_GWK".teco_cs_cw_e[1]
   //         State                  :="DB905_GWK".State[1]
END_REGION

REGION Network 9: Filling pump
         A     "DB009_Faults".Faults_Reset_FKT_M1;
         R     "DB822_Error_Tank".FeedPump[1].FLT_Dryrunsafety;
         R     "DB822_Error_Tank".FeedPump[1].FLT_Motorprotection;
         R     "DB822_Error_Tank".FeedPump[1].FLT_No_Barrel;
   //----- Störung Trockenlauf Befüllung
         A(;
         O     "K_Filling_Tank_C1";
         O     "K_Filling_Tank_C1_TL";
         );
         A     "DB702_Tank_Value".Tank[1].With_Filling_DryRun;
         L     s5t#5s;
         SD    "TM_Tank_Delay_DryRun_FeedPump_C1";
   //-
         A     "TM_Tank_Delay_DryRun_FeedPump_C1";
         AN    "S_DryRun_Feed_C1";
         AN    "DB822_Error_Tank".FeedPump[1].FLT_Dryrunsafety;
         S     "DB822_Error_Tank".FeedPump[1].FLT_Dryrunsafety;
         S     "DB009_Faults".Faults_FKT_Grp_3_M1;
         S     "DB009_Faults".Faultschanging_M1;
   //----- Störung Motorschutz Füllpumpe
   //    U     "F_FeedPump_C1"
   //    U     "DB702_Tank_Value".Tank[1].With_Filling_Pump
   //    UN    "DB822_Error_Tank".FeedPump[1].FLT_Motorprotection
   //    S     "DB822_Error_Tank".FeedPump[1].FLT_Motorprotection
   //    S     "DB009_Faults".Faults_FKT_Grp_3_M1
   //    S     "DB009_Faults".Faultschanging_M1
   //----- Störung Kein Fass vorhanden aber Befüllung angewählt
   //    U     "K_Filling_Tank_C1"
   //    UN    "S_BarrelDetection_C1"
   //    UN    "DB822_Error_Tank".FeedPump[1].FLT_No_Barrel
   //    S     "DB822_Error_Tank".FeedPump[1].FLT_No_Barrel
   //    S     "DB009_Faults".Faults_FKT_Grp_3_M1
   //    S     "DB009_Faults".Faultschanging_M1
   //----- Meldung Kein Fass vorhanden
   //    UN    "S_BarrelDetection_C1"
   //    UN    "DB822_Error_Tank".FeedPump[1].FLT_No_Barrel
         CLR;
         =     "DB822_Error_Tank".FeedPump[1].Mes_No_Barrel;
   //-----
         AN    "DB822_Error_Tank".FeedPump[1].FLT_No_Barrel;
         AN    "DB822_Error_Tank".FeedPump[1].Mes_No_Barrel;
         AN    "DB822_Error_Tank".FeedPump[1].FLT_Dryrunsafety;
         AN    "DB822_Error_Tank".FeedPump[1].FLT_Motorprotection;
         A     "DB702_Tank_Value".Tank[1].With_Filling_Pump;
         A(;
         O     "K_Filling_Tank_C1";
         O     "K_Filling_Tank_C1_TL";
         );

         =     "M_FeedPump_C1";
   //-----
END_REGION

REGION Network 10: Vacuum daytank
         CALL  "FC106_Vacuum"
         ( IN_Release           := "DB619_State_MPart".Operationmode[1].valid,
           IN_P_Vacuum          := "P_Vacuum_C1",
           IN_Timer_delay_Lock  := "TM_Vac1DelayLock",
           IN_Timer_delay_Pumpe := "TM_Vac1DelayPump",
           OUT_V_Lock_Vacuum    := "V_PressureVacuum_C1",
           OUT_V_Pump_Vacuum    := "V_PumpVacuum_C1",
           OUT_H_Vacuum_active  := #Temp_Vacuum_active,
           IO_Status            := "DB612_Tank_State".Vacuum[1]
         );
   //-----
END_REGION

